REGION Network 31
   RUNG wire#powerrail
      Contact( "SENSOR_DSBG_BASTIDOR_ABAJO_2" )
      Coil( "HMI_CUBA_FESTO".HMI_SENSOR_DSBG_BASTIDOR_ABAJO_2 )
   END_RUNG
   // the same network as SCL:
   "HMI_CUBA_FESTO".HMI_SENSOR_DSBG_BASTIDOR_ABAJO_2 := "SENSOR_DSBG_BASTIDOR_ABAJO_2";
END_REGION

REGION Network 32
   RUNG wire#powerrail
      Contact( "HMI_CUBA_FESTO".HMI_VALVULA_52_BIESTABLE_11 )
      S_Coil( "VALVULA_52_BIESTABLE_11" )
   END_RUNG
   RUNG wire#powerrail
      I_Contact( "HMI_CUBA_FESTO".HMI_VALVULA_52_BIESTABLE_11 )
      R_Coil( "VALVULA_52_BIESTABLE_11" )
   END_RUNG
   // the same network as SCL:
   IF "HMI_CUBA_FESTO".HMI_VALVULA_52_BIESTABLE_11 THEN "VALVULA_52_BIESTABLE_11" := TRUE; END_IF;
   IF NOT "HMI_CUBA_FESTO".HMI_VALVULA_52_BIESTABLE_11 THEN "VALVULA_52_BIESTABLE_11" := FALSE; END_IF;
END_REGION

REGION Network 33
   RUNG wire#powerrail
      Contact( "HMI_CUBA_FESTO".HMI_VALVULA_52_BIESTABLE_12 )
      S_Coil( "VALVULA_52_BIESTABLE_12" )
   END_RUNG
   RUNG wire#powerrail
      I_Contact( "HMI_CUBA_FESTO".HMI_VALVULA_52_BIESTABLE_12 )
      R_Coil( "VALVULA_52_BIESTABLE_12" )
   END_RUNG
   // the same network as SCL:
   IF "HMI_CUBA_FESTO".HMI_VALVULA_52_BIESTABLE_12 THEN "VALVULA_52_BIESTABLE_12" := TRUE; END_IF;
   IF NOT "HMI_CUBA_FESTO".HMI_VALVULA_52_BIESTABLE_12 THEN "VALVULA_52_BIESTABLE_12" := FALSE; END_IF;
END_REGION

REGION Network 34
   RUNG wire#powerrail
      Contact( "HMI_CUBA_FESTO".HMI_VALVULA_52_BIESTABLE_21 )
      S_Coil( "VALVULA_52_BIESTABLE_21" )
   END_RUNG
   RUNG wire#powerrail
      I_Contact( "HMI_CUBA_FESTO".HMI_VALVULA_52_BIESTABLE_21 )
      R_Coil( "VALVULA_52_BIESTABLE_21" )
   END_RUNG
   // the same network as SCL:
   IF "HMI_CUBA_FESTO".HMI_VALVULA_52_BIESTABLE_21 THEN "VALVULA_52_BIESTABLE_21" := TRUE; END_IF;
   IF NOT "HMI_CUBA_FESTO".HMI_VALVULA_52_BIESTABLE_21 THEN "VALVULA_52_BIESTABLE_21" := FALSE; END_IF;
END_REGION

REGION Network 35
   RUNG wire#powerrail
      Contact( "HMI_CUBA_FESTO".HMI_VALVULA_52_BIESTABLE_22 )
      S_Coil( "VALVULA_52_BIESTABLE_22" )
   END_RUNG
   RUNG wire#powerrail
      I_Contact( "HMI_CUBA_FESTO".HMI_VALVULA_52_BIESTABLE_22 )
      R_Coil( "VALVULA_52_BIESTABLE_22" )
   END_RUNG
   // the same network as SCL:
   IF "HMI_CUBA_FESTO".HMI_VALVULA_52_BIESTABLE_22 THEN "VALVULA_52_BIESTABLE_22" := TRUE; END_IF;
   IF NOT "HMI_CUBA_FESTO".HMI_VALVULA_52_BIESTABLE_22 THEN "VALVULA_52_BIESTABLE_22" := FALSE; END_IF;
END_REGION

REGION Network 36
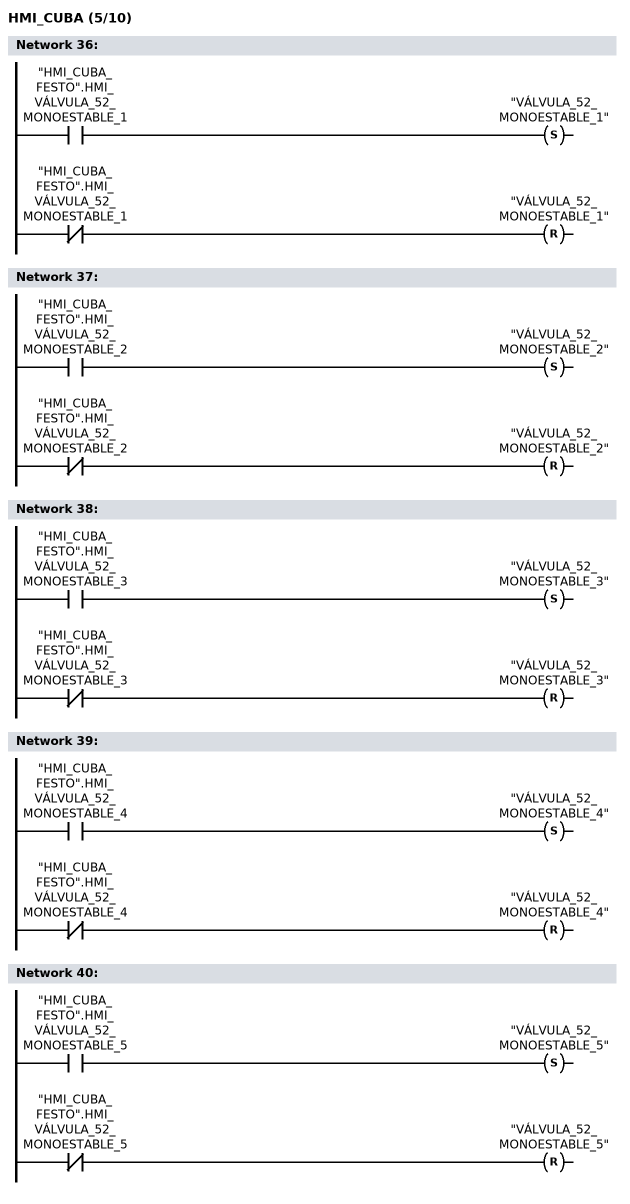
   RUNG wire#powerrail
      Contact( "HMI_CUBA_FESTO".HMI_VÁLVULA_52_MONOESTABLE_1 )
      S_Coil( "VÁLVULA_52_MONOESTABLE_1" )
   END_RUNG
   RUNG wire#powerrail
      I_Contact( "HMI_CUBA_FESTO".HMI_VÁLVULA_52_MONOESTABLE_1 )
      R_Coil( "VÁLVULA_52_MONOESTABLE_1" )
   END_RUNG
   // the same network as SCL:
   IF "HMI_CUBA_FESTO".HMI_VÁLVULA_52_MONOESTABLE_1 THEN "VÁLVULA_52_MONOESTABLE_1" := TRUE; END_IF;
   IF NOT "HMI_CUBA_FESTO".HMI_VÁLVULA_52_MONOESTABLE_1 THEN "VÁLVULA_52_MONOESTABLE_1" := FALSE; END_IF;
END_REGION

REGION Network 37
   RUNG wire#powerrail
      Contact( "HMI_CUBA_FESTO".HMI_VÁLVULA_52_MONOESTABLE_2 )
      S_Coil( "VÁLVULA_52_MONOESTABLE_2" )
   END_RUNG
   RUNG wire#powerrail
      I_Contact( "HMI_CUBA_FESTO".HMI_VÁLVULA_52_MONOESTABLE_2 )
      R_Coil( "VÁLVULA_52_MONOESTABLE_2" )
   END_RUNG
   // the same network as SCL:
   IF "HMI_CUBA_FESTO".HMI_VÁLVULA_52_MONOESTABLE_2 THEN "VÁLVULA_52_MONOESTABLE_2" := TRUE; END_IF;
   IF NOT "HMI_CUBA_FESTO".HMI_VÁLVULA_52_MONOESTABLE_2 THEN "VÁLVULA_52_MONOESTABLE_2" := FALSE; END_IF;
END_REGION

REGION Network 38
   RUNG wire#powerrail
      Contact( "HMI_CUBA_FESTO".HMI_VÁLVULA_52_MONOESTABLE_3 )
      S_Coil( "VÁLVULA_52_MONOESTABLE_3" )
   END_RUNG
   RUNG wire#powerrail
      I_Contact( "HMI_CUBA_FESTO".HMI_VÁLVULA_52_MONOESTABLE_3 )
      R_Coil( "VÁLVULA_52_MONOESTABLE_3" )
   END_RUNG
   // the same network as SCL:
   IF "HMI_CUBA_FESTO".HMI_VÁLVULA_52_MONOESTABLE_3 THEN "VÁLVULA_52_MONOESTABLE_3" := TRUE; END_IF;
   IF NOT "HMI_CUBA_FESTO".HMI_VÁLVULA_52_MONOESTABLE_3 THEN "VÁLVULA_52_MONOESTABLE_3" := FALSE; END_IF;
END_REGION

REGION Network 39
   RUNG wire#powerrail
      Contact( "HMI_CUBA_FESTO".HMI_VÁLVULA_52_MONOESTABLE_4 )
      S_Coil( "VÁLVULA_52_MONOESTABLE_4" )
   END_RUNG
   RUNG wire#powerrail
      I_Contact( "HMI_CUBA_FESTO".HMI_VÁLVULA_52_MONOESTABLE_4 )
      R_Coil( "VÁLVULA_52_MONOESTABLE_4" )
   END_RUNG
   // the same network as SCL:
   IF "HMI_CUBA_FESTO".HMI_VÁLVULA_52_MONOESTABLE_4 THEN "VÁLVULA_52_MONOESTABLE_4" := TRUE; END_IF;
   IF NOT "HMI_CUBA_FESTO".HMI_VÁLVULA_52_MONOESTABLE_4 THEN "VÁLVULA_52_MONOESTABLE_4" := FALSE; END_IF;
END_REGION

REGION Network 40
   RUNG wire#powerrail
      Contact( "HMI_CUBA_FESTO".HMI_VÁLVULA_52_MONOESTABLE_5 )
      S_Coil( "VÁLVULA_52_MONOESTABLE_5" )
   END_RUNG
   RUNG wire#powerrail
      I_Contact( "HMI_CUBA_FESTO".HMI_VÁLVULA_52_MONOESTABLE_5 )
      R_Coil( "VÁLVULA_52_MONOESTABLE_5" )
   END_RUNG
   // the same network as SCL:
   IF "HMI_CUBA_FESTO".HMI_VÁLVULA_52_MONOESTABLE_5 THEN "VÁLVULA_52_MONOESTABLE_5" := TRUE; END_IF;
   IF NOT "HMI_CUBA_FESTO".HMI_VÁLVULA_52_MONOESTABLE_5 THEN "VÁLVULA_52_MONOESTABLE_5" := FALSE; END_IF;
END_REGION

REGION Network 41
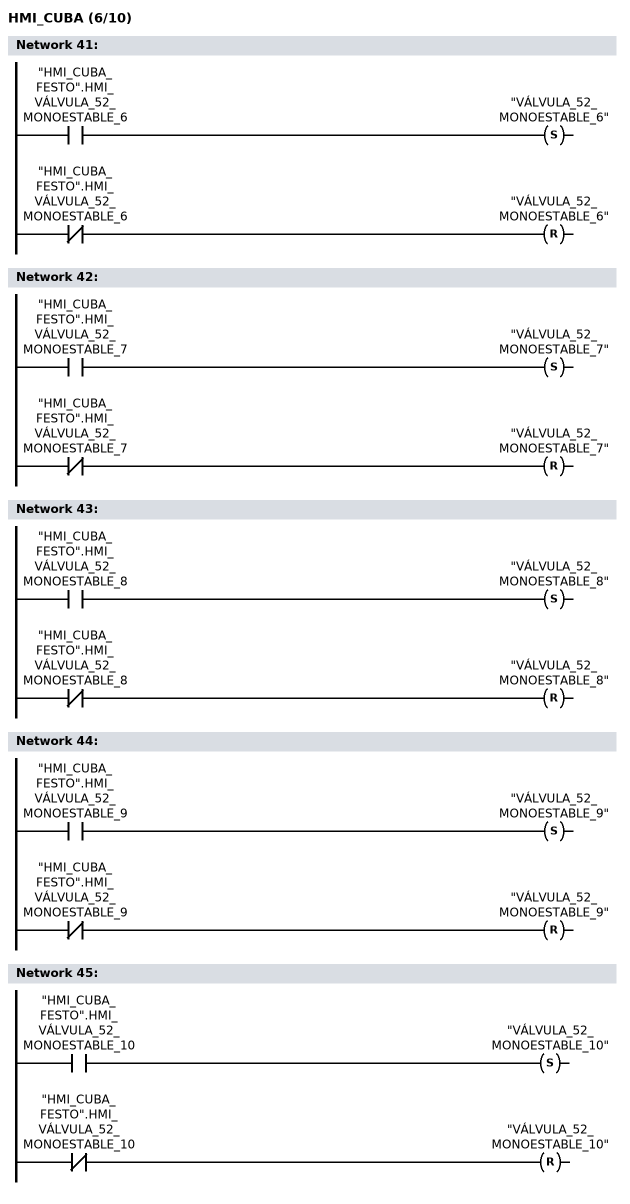
   RUNG wire#powerrail
      Contact( "HMI_CUBA_FESTO".HMI_VÁLVULA_52_MONOESTABLE_6 )
      S_Coil( "VÁLVULA_52_MONOESTABLE_6" )
   END_RUNG
   RUNG wire#powerrail
      I_Contact( "HMI_CUBA_FESTO".HMI_VÁLVULA_52_MONOESTABLE_6 )
      R_Coil( "VÁLVULA_52_MONOESTABLE_6" )
   END_RUNG
   // the same network as SCL:
   IF "HMI_CUBA_FESTO".HMI_VÁLVULA_52_MONOESTABLE_6 THEN "VÁLVULA_52_MONOESTABLE_6" := TRUE; END_IF;
   IF NOT "HMI_CUBA_FESTO".HMI_VÁLVULA_52_MONOESTABLE_6 THEN "VÁLVULA_52_MONOESTABLE_6" := FALSE; END_IF;
END_REGION

REGION Network 42
   RUNG wire#powerrail
      Contact( "HMI_CUBA_FESTO".HMI_VÁLVULA_52_MONOESTABLE_7 )
      S_Coil( "VÁLVULA_52_MONOESTABLE_7" )
   END_RUNG
   RUNG wire#powerrail
      I_Contact( "HMI_CUBA_FESTO".HMI_VÁLVULA_52_MONOESTABLE_7 )
      R_Coil( "VÁLVULA_52_MONOESTABLE_7" )
   END_RUNG
   // the same network as SCL:
   IF "HMI_CUBA_FESTO".HMI_VÁLVULA_52_MONOESTABLE_7 THEN "VÁLVULA_52_MONOESTABLE_7" := TRUE; END_IF;
   IF NOT "HMI_CUBA_FESTO".HMI_VÁLVULA_52_MONOESTABLE_7 THEN "VÁLVULA_52_MONOESTABLE_7" := FALSE; END_IF;
END_REGION

REGION Network 43
   RUNG wire#powerrail
      Contact( "HMI_CUBA_FESTO".HMI_VÁLVULA_52_MONOESTABLE_8 )
      S_Coil( "VÁLVULA_52_MONOESTABLE_8" )
   END_RUNG
   RUNG wire#powerrail
      I_Contact( "HMI_CUBA_FESTO".HMI_VÁLVULA_52_MONOESTABLE_8 )
      R_Coil( "VÁLVULA_52_MONOESTABLE_8" )
   END_RUNG
   // the same network as SCL:
   IF "HMI_CUBA_FESTO".HMI_VÁLVULA_52_MONOESTABLE_8 THEN "VÁLVULA_52_MONOESTABLE_8" := TRUE; END_IF;
   IF NOT "HMI_CUBA_FESTO".HMI_VÁLVULA_52_MONOESTABLE_8 THEN "VÁLVULA_52_MONOESTABLE_8" := FALSE; END_IF;
END_REGION

REGION Network 44
   RUNG wire#powerrail
      Contact( "HMI_CUBA_FESTO".HMI_VÁLVULA_52_MONOESTABLE_9 )
      S_Coil( "VÁLVULA_52_MONOESTABLE_9" )
   END_RUNG
   RUNG wire#powerrail
      I_Contact( "HMI_CUBA_FESTO".HMI_VÁLVULA_52_MONOESTABLE_9 )
      R_Coil( "VÁLVULA_52_MONOESTABLE_9" )
   END_RUNG
   // the same network as SCL:
   IF "HMI_CUBA_FESTO".HMI_VÁLVULA_52_MONOESTABLE_9 THEN "VÁLVULA_52_MONOESTABLE_9" := TRUE; END_IF;
   IF NOT "HMI_CUBA_FESTO".HMI_VÁLVULA_52_MONOESTABLE_9 THEN "VÁLVULA_52_MONOESTABLE_9" := FALSE; END_IF;
END_REGION

REGION Network 45
   RUNG wire#powerrail
      Contact( "HMI_CUBA_FESTO".HMI_VÁLVULA_52_MONOESTABLE_10 )
      S_Coil( "VÁLVULA_52_MONOESTABLE_10" )
   END_RUNG
   RUNG wire#powerrail
      I_Contact( "HMI_CUBA_FESTO".HMI_VÁLVULA_52_MONOESTABLE_10 )
      R_Coil( "VÁLVULA_52_MONOESTABLE_10" )
   END_RUNG
   // the same network as SCL:
   IF "HMI_CUBA_FESTO".HMI_VÁLVULA_52_MONOESTABLE_10 THEN "VÁLVULA_52_MONOESTABLE_10" := TRUE; END_IF;
   IF NOT "HMI_CUBA_FESTO".HMI_VÁLVULA_52_MONOESTABLE_10 THEN "VÁLVULA_52_MONOESTABLE_10" := FALSE; END_IF;
END_REGION

REGION Network 46
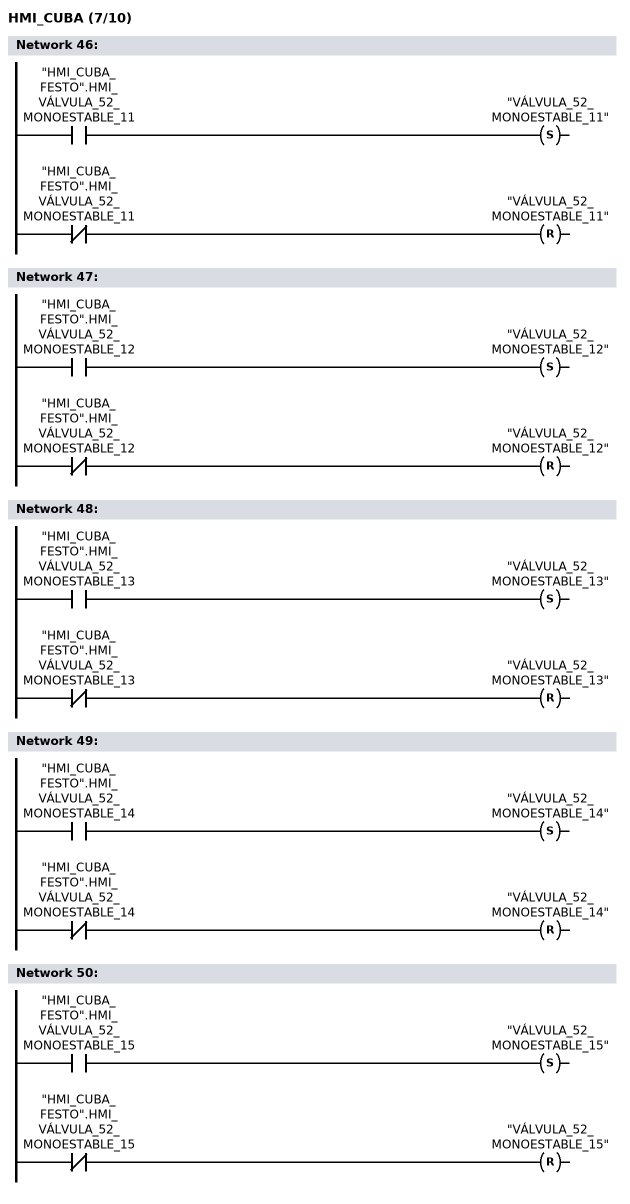
   RUNG wire#powerrail
      Contact( "HMI_CUBA_FESTO".HMI_VÁLVULA_52_MONOESTABLE_11 )
      S_Coil( "VÁLVULA_52_MONOESTABLE_11" )
   END_RUNG
   RUNG wire#powerrail
      I_Contact( "HMI_CUBA_FESTO".HMI_VÁLVULA_52_MONOESTABLE_11 )
      R_Coil( "VÁLVULA_52_MONOESTABLE_11" )
   END_RUNG
   // the same network as SCL:
   IF "HMI_CUBA_FESTO".HMI_VÁLVULA_52_MONOESTABLE_11 THEN "VÁLVULA_52_MONOESTABLE_11" := TRUE; END_IF;
   IF NOT "HMI_CUBA_FESTO".HMI_VÁLVULA_52_MONOESTABLE_11 THEN "VÁLVULA_52_MONOESTABLE_11" := FALSE; END_IF;
END_REGION

REGION Network 47
   RUNG wire#powerrail
      Contact( "HMI_CUBA_FESTO".HMI_VÁLVULA_52_MONOESTABLE_12 )
      S_Coil( "VÁLVULA_52_MONOESTABLE_12" )
   END_RUNG
   RUNG wire#powerrail
      I_Contact( "HMI_CUBA_FESTO".HMI_VÁLVULA_52_MONOESTABLE_12 )
      R_Coil( "VÁLVULA_52_MONOESTABLE_12" )
   END_RUNG
   // the same network as SCL:
   IF "HMI_CUBA_FESTO".HMI_VÁLVULA_52_MONOESTABLE_12 THEN "VÁLVULA_52_MONOESTABLE_12" := TRUE; END_IF;
   IF NOT "HMI_CUBA_FESTO".HMI_VÁLVULA_52_MONOESTABLE_12 THEN "VÁLVULA_52_MONOESTABLE_12" := FALSE; END_IF;
END_REGION

REGION Network 48
   RUNG wire#powerrail
      Contact( "HMI_CUBA_FESTO".HMI_VÁLVULA_52_MONOESTABLE_13 )
      S_Coil( "VÁLVULA_52_MONOESTABLE_13" )
   END_RUNG
   RUNG wire#powerrail
      I_Contact( "HMI_CUBA_FESTO".HMI_VÁLVULA_52_MONOESTABLE_13 )
      R_Coil( "VÁLVULA_52_MONOESTABLE_13" )
   END_RUNG
   // the same network as SCL:
   IF "HMI_CUBA_FESTO".HMI_VÁLVULA_52_MONOESTABLE_13 THEN "VÁLVULA_52_MONOESTABLE_13" := TRUE; END_IF;
   IF NOT "HMI_CUBA_FESTO".HMI_VÁLVULA_52_MONOESTABLE_13 THEN "VÁLVULA_52_MONOESTABLE_13" := FALSE; END_IF;
END_REGION

REGION Network 49
   RUNG wire#powerrail
      Contact( "HMI_CUBA_FESTO".HMI_VÁLVULA_52_MONOESTABLE_14 )
      S_Coil( "VÁLVULA_52_MONOESTABLE_14" )
   END_RUNG
   RUNG wire#powerrail
      I_Contact( "HMI_CUBA_FESTO".HMI_VÁLVULA_52_MONOESTABLE_14 )
      R_Coil( "VÁLVULA_52_MONOESTABLE_14" )
   END_RUNG
   // the same network as SCL:
   IF "HMI_CUBA_FESTO".HMI_VÁLVULA_52_MONOESTABLE_14 THEN "VÁLVULA_52_MONOESTABLE_14" := TRUE; END_IF;
   IF NOT "HMI_CUBA_FESTO".HMI_VÁLVULA_52_MONOESTABLE_14 THEN "VÁLVULA_52_MONOESTABLE_14" := FALSE; END_IF;
END_REGION

REGION Network 50
   RUNG wire#powerrail
      Contact( "HMI_CUBA_FESTO".HMI_VÁLVULA_52_MONOESTABLE_15 )
      S_Coil( "VÁLVULA_52_MONOESTABLE_15" )
   END_RUNG
   RUNG wire#powerrail
      I_Contact( "HMI_CUBA_FESTO".HMI_VÁLVULA_52_MONOESTABLE_15 )
      R_Coil( "VÁLVULA_52_MONOESTABLE_15" )
   END_RUNG
   // the same network as SCL:
   IF "HMI_CUBA_FESTO".HMI_VÁLVULA_52_MONOESTABLE_15 THEN "VÁLVULA_52_MONOESTABLE_15" := TRUE; END_IF;
   IF NOT "HMI_CUBA_FESTO".HMI_VÁLVULA_52_MONOESTABLE_15 THEN "VÁLVULA_52_MONOESTABLE_15" := FALSE; END_IF;
END_REGION

REGION Network 51
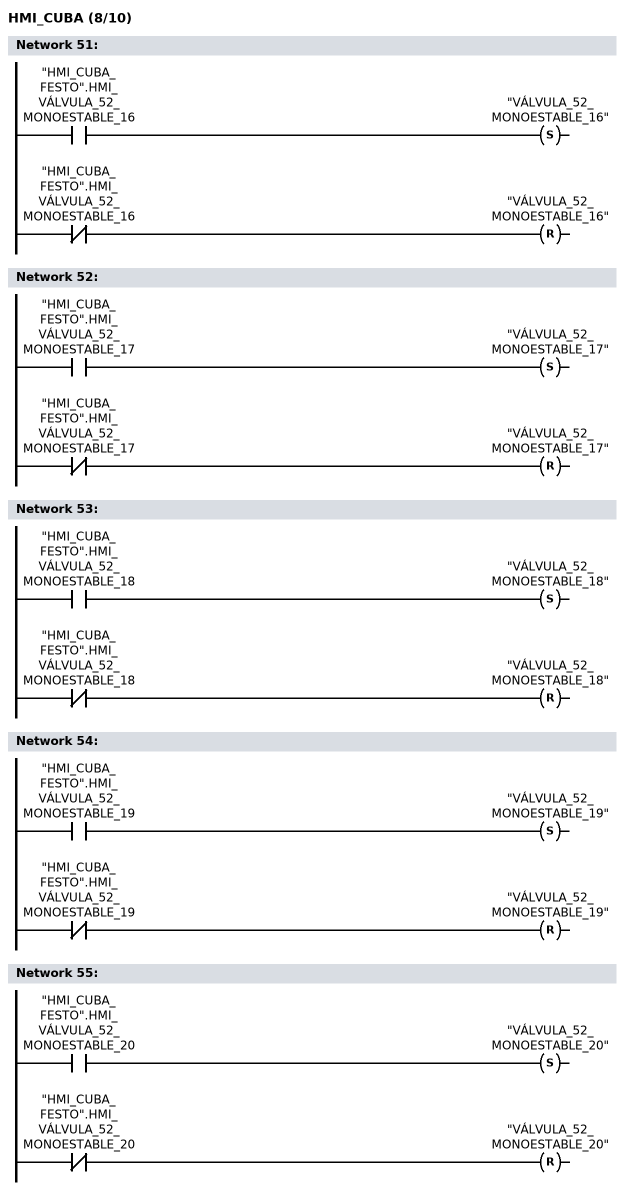
   RUNG wire#powerrail
      Contact( "HMI_CUBA_FESTO".HMI_VÁLVULA_52_MONOESTABLE_16 )
      S_Coil( "VÁLVULA_52_MONOESTABLE_16" )
   END_RUNG
   RUNG wire#powerrail
      I_Contact( "HMI_CUBA_FESTO".HMI_VÁLVULA_52_MONOESTABLE_16 )
      R_Coil( "VÁLVULA_52_MONOESTABLE_16" )
   END_RUNG
   // the same network as SCL:
   IF "HMI_CUBA_FESTO".HMI_VÁLVULA_52_MONOESTABLE_16 THEN "VÁLVULA_52_MONOESTABLE_16" := TRUE; END_IF;
   IF NOT "HMI_CUBA_FESTO".HMI_VÁLVULA_52_MONOESTABLE_16 THEN "VÁLVULA_52_MONOESTABLE_16" := FALSE; END_IF;
END_REGION

REGION Network 52
   RUNG wire#powerrail
      Contact( "HMI_CUBA_FESTO".HMI_VÁLVULA_52_MONOESTABLE_17 )
      S_Coil( "VÁLVULA_52_MONOESTABLE_17" )
   END_RUNG
   RUNG wire#powerrail
      I_Contact( "HMI_CUBA_FESTO".HMI_VÁLVULA_52_MONOESTABLE_17 )
      R_Coil( "VÁLVULA_52_MONOESTABLE_17" )
   END_RUNG
   // the same network as SCL:
   IF "HMI_CUBA_FESTO".HMI_VÁLVULA_52_MONOESTABLE_17 THEN "VÁLVULA_52_MONOESTABLE_17" := TRUE; END_IF;
   IF NOT "HMI_CUBA_FESTO".HMI_VÁLVULA_52_MONOESTABLE_17 THEN "VÁLVULA_52_MONOESTABLE_17" := FALSE; END_IF;
END_REGION

REGION Network 53
   RUNG wire#powerrail
      Contact( "HMI_CUBA_FESTO".HMI_VÁLVULA_52_MONOESTABLE_18 )
      S_Coil( "VÁLVULA_52_MONOESTABLE_18" )
   END_RUNG
   RUNG wire#powerrail
      I_Contact( "HMI_CUBA_FESTO".HMI_VÁLVULA_52_MONOESTABLE_18 )
      R_Coil( "VÁLVULA_52_MONOESTABLE_18" )
   END_RUNG
   // the same network as SCL:
   IF "HMI_CUBA_FESTO".HMI_VÁLVULA_52_MONOESTABLE_18 THEN "VÁLVULA_52_MONOESTABLE_18" := TRUE; END_IF;
   IF NOT "HMI_CUBA_FESTO".HMI_VÁLVULA_52_MONOESTABLE_18 THEN "VÁLVULA_52_MONOESTABLE_18" := FALSE; END_IF;
END_REGION

REGION Network 54
   RUNG wire#powerrail
      Contact( "HMI_CUBA_FESTO".HMI_VÁLVULA_52_MONOESTABLE_19 )
      S_Coil( "VÁLVULA_52_MONOESTABLE_19" )
   END_RUNG
   RUNG wire#powerrail
      I_Contact( "HMI_CUBA_FESTO".HMI_VÁLVULA_52_MONOESTABLE_19 )
      R_Coil( "VÁLVULA_52_MONOESTABLE_19" )
   END_RUNG
   // the same network as SCL:
   IF "HMI_CUBA_FESTO".HMI_VÁLVULA_52_MONOESTABLE_19 THEN "VÁLVULA_52_MONOESTABLE_19" := TRUE; END_IF;
   IF NOT "HMI_CUBA_FESTO".HMI_VÁLVULA_52_MONOESTABLE_19 THEN "VÁLVULA_52_MONOESTABLE_19" := FALSE; END_IF;
END_REGION

REGION Network 55
   RUNG wire#powerrail
      Contact( "HMI_CUBA_FESTO".HMI_VÁLVULA_52_MONOESTABLE_20 )
      S_Coil( "VÁLVULA_52_MONOESTABLE_20" )
   END_RUNG
   RUNG wire#powerrail
      I_Contact( "HMI_CUBA_FESTO".HMI_VÁLVULA_52_MONOESTABLE_20 )
      R_Coil( "VÁLVULA_52_MONOESTABLE_20" )
   END_RUNG
   // the same network as SCL:
   IF "HMI_CUBA_FESTO".HMI_VÁLVULA_52_MONOESTABLE_20 THEN "VÁLVULA_52_MONOESTABLE_20" := TRUE; END_IF;
   IF NOT "HMI_CUBA_FESTO".HMI_VÁLVULA_52_MONOESTABLE_20 THEN "VÁLVULA_52_MONOESTABLE_20" := FALSE; END_IF;
END_REGION

REGION Network 56
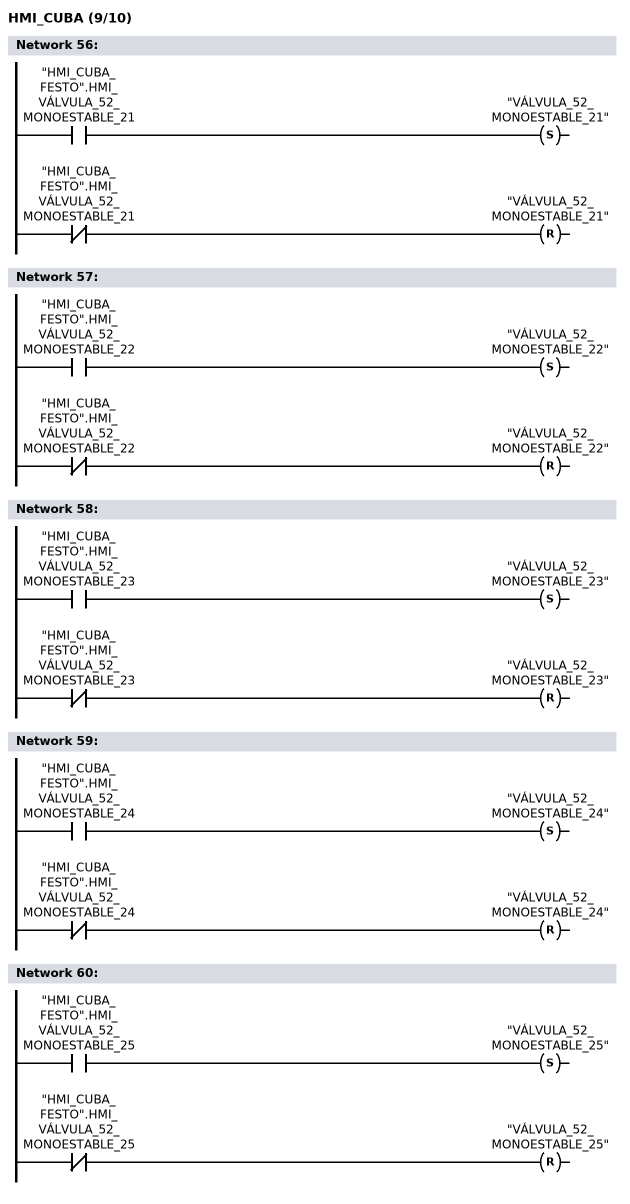
   RUNG wire#powerrail
      Contact( "HMI_CUBA_FESTO".HMI_VÁLVULA_52_MONOESTABLE_21 )
      S_Coil( "VÁLVULA_52_MONOESTABLE_21" )
   END_RUNG
   RUNG wire#powerrail
      I_Contact( "HMI_CUBA_FESTO".HMI_VÁLVULA_52_MONOESTABLE_21 )
      R_Coil( "VÁLVULA_52_MONOESTABLE_21" )
   END_RUNG
   // the same network as SCL:
   IF "HMI_CUBA_FESTO".HMI_VÁLVULA_52_MONOESTABLE_21 THEN "VÁLVULA_52_MONOESTABLE_21" := TRUE; END_IF;
   IF NOT "HMI_CUBA_FESTO".HMI_VÁLVULA_52_MONOESTABLE_21 THEN "VÁLVULA_52_MONOESTABLE_21" := FALSE; END_IF;
END_REGION

REGION Network 57
   RUNG wire#powerrail
      Contact( "HMI_CUBA_FESTO".HMI_VÁLVULA_52_MONOESTABLE_22 )
      S_Coil( "VÁLVULA_52_MONOESTABLE_22" )
   END_RUNG
   RUNG wire#powerrail
      I_Contact( "HMI_CUBA_FESTO".HMI_VÁLVULA_52_MONOESTABLE_22 )
      R_Coil( "VÁLVULA_52_MONOESTABLE_22" )
   END_RUNG
   // the same network as SCL:
   IF "HMI_CUBA_FESTO".HMI_VÁLVULA_52_MONOESTABLE_22 THEN "VÁLVULA_52_MONOESTABLE_22" := TRUE; END_IF;
   IF NOT "HMI_CUBA_FESTO".HMI_VÁLVULA_52_MONOESTABLE_22 THEN "VÁLVULA_52_MONOESTABLE_22" := FALSE; END_IF;
END_REGION

REGION Network 58
   RUNG wire#powerrail
      Contact( "HMI_CUBA_FESTO".HMI_VÁLVULA_52_MONOESTABLE_23 )
      S_Coil( "VÁLVULA_52_MONOESTABLE_23" )
   END_RUNG
   RUNG wire#powerrail
      I_Contact( "HMI_CUBA_FESTO".HMI_VÁLVULA_52_MONOESTABLE_23 )
      R_Coil( "VÁLVULA_52_MONOESTABLE_23" )
   END_RUNG
   // the same network as SCL:
   IF "HMI_CUBA_FESTO".HMI_VÁLVULA_52_MONOESTABLE_23 THEN "VÁLVULA_52_MONOESTABLE_23" := TRUE; END_IF;
   IF NOT "HMI_CUBA_FESTO".HMI_VÁLVULA_52_MONOESTABLE_23 THEN "VÁLVULA_52_MONOESTABLE_23" := FALSE; END_IF;
END_REGION

REGION Network 59
   RUNG wire#powerrail
      Contact( "HMI_CUBA_FESTO".HMI_VÁLVULA_52_MONOESTABLE_24 )
      S_Coil( "VÁLVULA_52_MONOESTABLE_24" )
   END_RUNG
   RUNG wire#powerrail
      I_Contact( "HMI_CUBA_FESTO".HMI_VÁLVULA_52_MONOESTABLE_24 )
      R_Coil( "VÁLVULA_52_MONOESTABLE_24" )
   END_RUNG
   // the same network as SCL:
   IF "HMI_CUBA_FESTO".HMI_VÁLVULA_52_MONOESTABLE_24 THEN "VÁLVULA_52_MONOESTABLE_24" := TRUE; END_IF;
   IF NOT "HMI_CUBA_FESTO".HMI_VÁLVULA_52_MONOESTABLE_24 THEN "VÁLVULA_52_MONOESTABLE_24" := FALSE; END_IF;
END_REGION

REGION Network 60
   RUNG wire#powerrail
      Contact( "HMI_CUBA_FESTO".HMI_VÁLVULA_52_MONOESTABLE_25 )
      S_Coil( "VÁLVULA_52_MONOESTABLE_25" )
   END_RUNG
   RUNG wire#powerrail
      I_Contact( "HMI_CUBA_FESTO".HMI_VÁLVULA_52_MONOESTABLE_25 )
      R_Coil( "VÁLVULA_52_MONOESTABLE_25" )
   END_RUNG
   // the same network as SCL:
   IF "HMI_CUBA_FESTO".HMI_VÁLVULA_52_MONOESTABLE_25 THEN "VÁLVULA_52_MONOESTABLE_25" := TRUE; END_IF;
   IF NOT "HMI_CUBA_FESTO".HMI_VÁLVULA_52_MONOESTABLE_25 THEN "VÁLVULA_52_MONOESTABLE_25" := FALSE; END_IF;
END_REGION

REGION Network 61
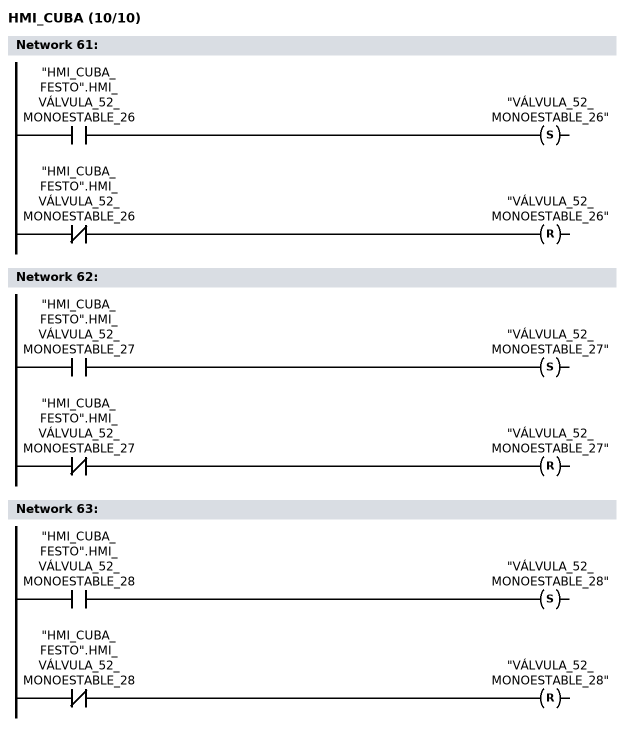
   RUNG wire#powerrail
      Contact( "HMI_CUBA_FESTO".HMI_VÁLVULA_52_MONOESTABLE_26 )
      S_Coil( "VÁLVULA_52_MONOESTABLE_26" )
   END_RUNG
   RUNG wire#powerrail
      I_Contact( "HMI_CUBA_FESTO".HMI_VÁLVULA_52_MONOESTABLE_26 )
      R_Coil( "VÁLVULA_52_MONOESTABLE_26" )
   END_RUNG
   // the same network as SCL:
   IF "HMI_CUBA_FESTO".HMI_VÁLVULA_52_MONOESTABLE_26 THEN "VÁLVULA_52_MONOESTABLE_26" := TRUE; END_IF;
   IF NOT "HMI_CUBA_FESTO".HMI_VÁLVULA_52_MONOESTABLE_26 THEN "VÁLVULA_52_MONOESTABLE_26" := FALSE; END_IF;
END_REGION

REGION Network 62
   RUNG wire#powerrail
      Contact( "HMI_CUBA_FESTO".HMI_VÁLVULA_52_MONOESTABLE_27 )
      S_Coil( "VÁLVULA_52_MONOESTABLE_27" )
   END_RUNG
   RUNG wire#powerrail
      I_Contact( "HMI_CUBA_FESTO".HMI_VÁLVULA_52_MONOESTABLE_27 )
      R_Coil( "VÁLVULA_52_MONOESTABLE_27" )
   END_RUNG
   // the same network as SCL:
   IF "HMI_CUBA_FESTO".HMI_VÁLVULA_52_MONOESTABLE_27 THEN "VÁLVULA_52_MONOESTABLE_27" := TRUE; END_IF;
   IF NOT "HMI_CUBA_FESTO".HMI_VÁLVULA_52_MONOESTABLE_27 THEN "VÁLVULA_52_MONOESTABLE_27" := FALSE; END_IF;
END_REGION

REGION Network 63
   RUNG wire#powerrail
      Contact( "HMI_CUBA_FESTO".HMI_VÁLVULA_52_MONOESTABLE_28 )
      S_Coil( "VÁLVULA_52_MONOESTABLE_28" )
   END_RUNG
   RUNG wire#powerrail
      I_Contact( "HMI_CUBA_FESTO".HMI_VÁLVULA_52_MONOESTABLE_28 )
      R_Coil( "VÁLVULA_52_MONOESTABLE_28" )
   END_RUNG
   // the same network as SCL:
   IF "HMI_CUBA_FESTO".HMI_VÁLVULA_52_MONOESTABLE_28 THEN "VÁLVULA_52_MONOESTABLE_28" := TRUE; END_IF;
   IF NOT "HMI_CUBA_FESTO".HMI_VÁLVULA_52_MONOESTABLE_28 THEN "VÁLVULA_52_MONOESTABLE_28" := FALSE; END_IF;
END_REGION
END_FUNCTION_BLOCK

FUNCTION_BLOCK "GIRO_POSITIVO"   // FB10, LAD
{ S7_Optimized_Access := 'TRUE' }
VERSION : 0.1
   VAR_TEMP   // added for the SCL form of the ladder/FBD networks
      _w1 : Bool;
   END_VAR
BEGIN

REGION Network 1: Estado 1
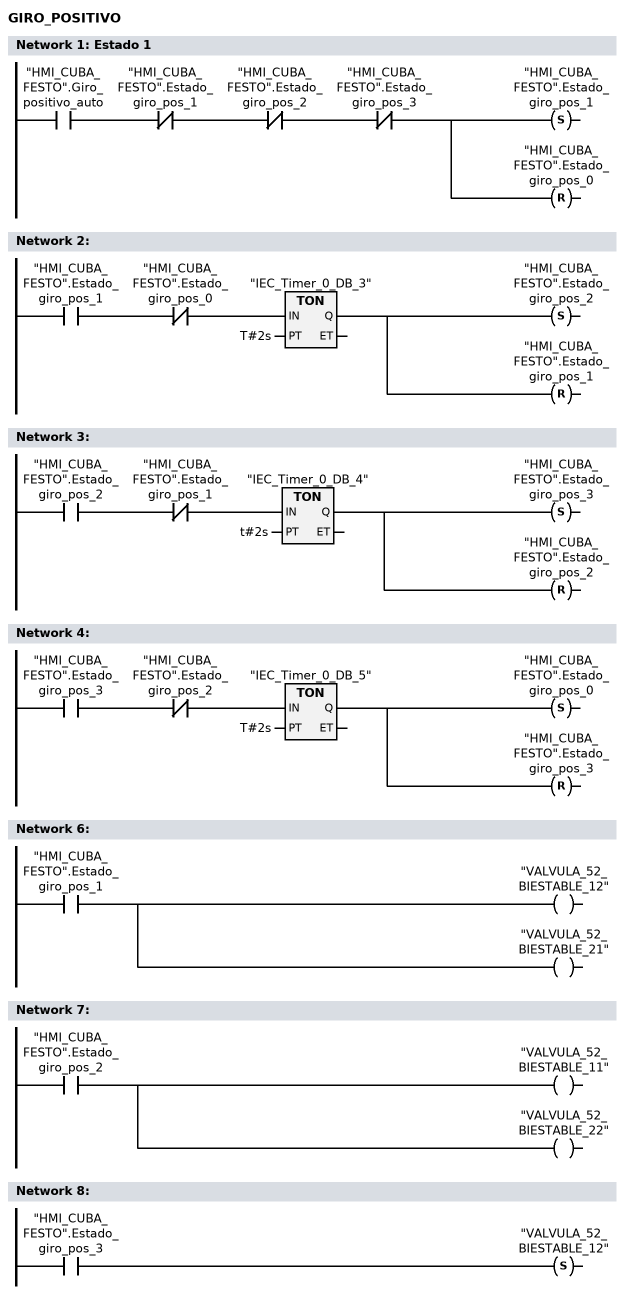
   RUNG wire#powerrail
      Contact( "HMI_CUBA_FESTO".Giro_positivo_auto )
      I_Contact( "HMI_CUBA_FESTO".Estado_giro_pos_1 )
      I_Contact( "HMI_CUBA_FESTO".Estado_giro_pos_2 )
      I_Contact( "HMI_CUBA_FESTO".Estado_giro_pos_3 )
      wire#w1
      S_Coil( "HMI_CUBA_FESTO".Estado_giro_pos_1 )
   END_RUNG
   RUNG wire#w1
      R_Coil( "HMI_CUBA_FESTO".Estado_giro_pos_0 )
   END_RUNG
   // the same network as SCL:
   #_w1 := "HMI_CUBA_FESTO".Giro_positivo_auto AND NOT "HMI_CUBA_FESTO".Estado_giro_pos_1 AND NOT "HMI_CUBA_FESTO".Estado_giro_pos_2 AND NOT "HMI_CUBA_FESTO".Estado_giro_pos_3;
   IF #_w1 THEN
       "HMI_CUBA_FESTO".Estado_giro_pos_1 := TRUE;
       "HMI_CUBA_FESTO".Estado_giro_pos_0 := FALSE;
   END_IF;
END_REGION

REGION Network 2
   "IEC_Timer_0_DB_3".TON(IN := "HMI_CUBA_FESTO".Estado_giro_pos_1 AND NOT "HMI_CUBA_FESTO".Estado_giro_pos_0,
                          PT := T#2s);
   IF "IEC_Timer_0_DB_3".Q THEN
       "HMI_CUBA_FESTO".Estado_giro_pos_2 := TRUE;
       "HMI_CUBA_FESTO".Estado_giro_pos_1 := FALSE;
   END_IF;
END_REGION

REGION Network 3
   "IEC_Timer_0_DB_4".TON(IN := "HMI_CUBA_FESTO".Estado_giro_pos_2 AND NOT "HMI_CUBA_FESTO".Estado_giro_pos_1,
                          PT := t#2s);
   IF "IEC_Timer_0_DB_4".Q THEN
       "HMI_CUBA_FESTO".Estado_giro_pos_3 := TRUE;
       "HMI_CUBA_FESTO".Estado_giro_pos_2 := FALSE;
   END_IF;
END_REGION

REGION Network 4
   "IEC_Timer_0_DB_5".TON(IN := "HMI_CUBA_FESTO".Estado_giro_pos_3 AND NOT "HMI_CUBA_FESTO".Estado_giro_pos_2,
                          PT := T#2s);
   IF "IEC_Timer_0_DB_5".Q THEN
       "HMI_CUBA_FESTO".Estado_giro_pos_0 := TRUE;
       "HMI_CUBA_FESTO".Estado_giro_pos_3 := FALSE;
   END_IF;
END_REGION

REGION Network 6
   RUNG wire#powerrail
      Contact( "HMI_CUBA_FESTO".Estado_giro_pos_1 )
      wire#w1
      Coil( "VALVULA_52_BIESTABLE_12" )
   END_RUNG
   RUNG wire#w1
      Coil( "VALVULA_52_BIESTABLE_21" )
   END_RUNG
   // the same network as SCL:
   "VALVULA_52_BIESTABLE_12" := "HMI_CUBA_FESTO".Estado_giro_pos_1;
   "VALVULA_52_BIESTABLE_21" := "HMI_CUBA_FESTO".Estado_giro_pos_1;
END_REGION

REGION Network 7
   RUNG wire#powerrail
      Contact( "HMI_CUBA_FESTO".Estado_giro_pos_2 )
      wire#w1
      Coil( "VALVULA_52_BIESTABLE_11" )
   END_RUNG
   RUNG wire#w1
      Coil( "VALVULA_52_BIESTABLE_22" )
   END_RUNG
   // the same network as SCL:
   "VALVULA_52_BIESTABLE_11" := "HMI_CUBA_FESTO".Estado_giro_pos_2;
   "VALVULA_52_BIESTABLE_22" := "HMI_CUBA_FESTO".Estado_giro_pos_2;
END_REGION

REGION Network 8
   RUNG wire#powerrail
      Contact( "HMI_CUBA_FESTO".Estado_giro_pos_3 )
      S_Coil( "VALVULA_52_BIESTABLE_12" )
   END_RUNG
   // the same network as SCL:
   IF "HMI_CUBA_FESTO".Estado_giro_pos_3 THEN "VALVULA_52_BIESTABLE_12" := TRUE; END_IF;
END_REGION
END_FUNCTION_BLOCK

FUNCTION_BLOCK "GIRO_NEGATIVO_1"   // FB14, LAD
{ S7_Optimized_Access := 'TRUE' }
VERSION : 0.1
   VAR_TEMP   // added for the SCL form of the ladder/FBD networks
      _w1 : Bool;
   END_VAR
BEGIN

REGION Network 1: Estado 1